(* Logix 5000 project; controller MV vendor 1 type 14 code 217 rev 31.11; software revision 31.00; part 51 of 53 *)
(* tags used below, declared in another part *)
   Alarm_Reset : BOOL;
   CWD : CHECKWORD_FLAGS;
   Default_Check_Time : DINT;
   Item_Faults_Are_Latched : BOOL;
   Item_Simulation_Flag : BOOL;
   MV_MV10R : PlantItem;   // MV10R
   MV_MV10R_ALARM : ALARM_DIGITAL;
   MV_MV10R_D : ALIAS FOR Remote_IO:13:O.Data.9;   // Rouser drive MV10
   MV_MV10R_R : ALIAS FOR Remote_IO:15:I.Data.9;   // MV10 Rouser running signal
   MV_MV11R : PlantItem;   // MV11R
   MV_MV11R_ALARM : ALARM_DIGITAL;
   MV_MV11R_D : ALIAS FOR Remote_IO:13:O.Data.10;   // Rouser drive MV11
   MV_MV11R_R : ALIAS FOR Remote_IO:15:I.Data.10;   // MV11 Rouser running signal
   MV_MV12R : PlantItem;   // MV12R
   MV_MV12R_ALARM : ALARM_DIGITAL;
   MV_MV12R_D : ALIAS FOR Remote_IO:13:O.Data.11;   // Rouser drive MV12
   MV_MV12R_R : ALIAS FOR Remote_IO:15:I.Data.11;   // MV12 Rouser running signal
   MV_MV13R : PlantItem;   // MV13R
   MV_MV13R_ALARM : ALARM_DIGITAL;
   MV_MV13R_D : ALIAS FOR Remote_IO:13:O.Data.12;   // Rouser drive MV13
   MV_MV13R_R : ALIAS FOR Remote_IO:15:I.Data.12;   // MV13 Rouser running signal
   MV_MV14R : PlantItem;   // MV14R
   MV_MV14R_ALARM : ALARM_DIGITAL;
   MV_MV14R_D : ALIAS FOR Remote_IO:13:O.Data.13;   // Rouser drive MV14
   MV_MV14R_R : ALIAS FOR Remote_IO:15:I.Data.13;   // MV14 Rouser running signal
   MV_MV15R : PlantItem;   // MV15R
   MV_MV15R_ALARM : ALARM_DIGITAL;
   MV_MV15R_D : ALIAS FOR Remote_IO:13:O.Data.14;   // Rouser drive MV15
   MV_MV15R_R : ALIAS FOR Remote_IO:15:I.Data.14;   // MV15 Rouser running signal
   MV_MV16R : PlantItem;   // MV16R
   MV_MV16R_ALARM : ALARM_DIGITAL;
   MV_MV16R_D : ALIAS FOR Remote_IO:13:O.Data.15;   // Rouser drive MV16
   MV_MV16R_R : ALIAS FOR Remote_IO:15:I.Data.15;   // MV16 Rouser running signal
   MV_MV17R : PlantItem;   // MV17R
   MV_MV17R_ALARM : ALARM_DIGITAL;
   MV_MV17R_D : ALIAS FOR Remote_IO:14:O.Data.0;   // Rouser drive MV17
   MV_MV17R_R : ALIAS FOR Remote_IO:15:I.Data.16;   // MV17 Rouser running signal
   MV_MV18R : PlantItem;   // MV18R
   MV_MV18R_ALARM : ALARM_DIGITAL;
   MV_MV18R_D : ALIAS FOR Remote_IO:14:O.Data.1;
   MV_MV18R_R : ALIAS FOR Remote_IO:15:I.Data.17;   // MV18 Rouser running signal
   MV_MV19R : PlantItem;   // MV19R
   MV_MV19R_ALARM : ALARM_DIGITAL;
   MV_MV19R_D : ALIAS FOR Remote_IO:14:O.Data.2;   // Rouser drive MV19
   MV_MV19R_R : ALIAS FOR Remote_IO:15:I.Data.18;   // MV19 Rouser running signal
   MV_MV1R : PlantItem;   // MV1R
   MV_MV1R_ALARM : ALARM_DIGITAL;
   MV_MV1R_D : ALIAS FOR Remote_IO:13:O.Data.0;   // Rouser drive MV1
   MV_MV1R_R : ALIAS FOR Remote_IO:15:I.Data.0;
   MV_MV2R : PlantItem;   // MV2R
   MV_MV2R_ALARM : ALARM_DIGITAL;
   MV_MV2R_D : ALIAS FOR Remote_IO:13:O.Data.1;
   MV_MV2R_R : ALIAS FOR Remote_IO:15:I.Data.1;   // MV2 Rouser running signal
   MV_MV30R : PlantItem;   // MV30R
   MV_MV30R_ALARM : ALARM_DIGITAL;
   MV_MV30R_D : ALIAS FOR Remote_IO:14:O.Data.3;   // Rouser drive MV30
   MV_MV30R_R : ALIAS FOR Remote_IO:15:I.Data.19;   // MV30 Rouser running signal
   MV_MV31R : PlantItem;   // MV31R
   MV_MV31R_ALARM : ALARM_DIGITAL;
   MV_MV31R_D : ALIAS FOR Remote_IO:14:O.Data.4;   // Rouser drive MV31
   MV_MV31R_R : ALIAS FOR Remote_IO:15:I.Data.20;   // MV31 Rouser running signal
   MV_MV32R : PlantItem;   // MV32R
   MV_MV32R_ALARM : ALARM_DIGITAL;
   MV_MV32R_D : ALIAS FOR Remote_IO:14:O.Data.5;   // Rouser drive MV32
   MV_MV32R_R : ALIAS FOR Remote_IO:15:I.Data.21;   // MV32 Rouser running signal
   MV_MV33R : PlantItem;   // MV33R
   MV_MV33R_ALARM : ALARM_DIGITAL;
   MV_MV33R_D : ALIAS FOR Remote_IO:14:O.Data.6;   // Rouser drive MV33
   MV_MV33R_R : ALIAS FOR Remote_IO:15:I.Data.22;   // MV33 Rouser running signal
   MV_MV34R : PlantItem;   // MV34R
   MV_MV34R_ALARM : ALARM_DIGITAL;
   MV_MV34R_D : ALIAS FOR Remote_IO:14:O.Data.7;   // Rouser drive MV34
   MV_MV34R_R : ALIAS FOR Remote_IO:15:I.Data.23;   // MV34 Rouser running signal
   MV_MV3R : PlantItem;   // MV3R
   MV_MV3R_ALARM : ALARM_DIGITAL;
   MV_MV3R_D : ALIAS FOR Remote_IO:13:O.Data.2;   // Rouser drive MV3
   MV_MV3R_R : ALIAS FOR Remote_IO:15:I.Data.2;   // MV3 Rouser running signal
   MV_MV4R : PlantItem;   // MV4R
   MV_MV4R_ALARM : ALARM_DIGITAL;
   MV_MV4R_D : ALIAS FOR Remote_IO:13:O.Data.3;   // Rouser drive MV4
   MV_MV4R_R : ALIAS FOR Remote_IO:15:I.Data.3;   // MV4 Rouser running signal
   MV_MV5R : PlantItem;   // MV5R
   MV_MV5R_ALARM : ALARM_DIGITAL;
   MV_MV5R_D : ALIAS FOR Remote_IO:13:O.Data.4;   // Rouser drive MV5
   MV_MV5R_R : ALIAS FOR Remote_IO:15:I.Data.4;   // MV5 Rouser running signal
   MV_MV6R : PlantItem;   // MV6R
   MV_MV6R_ALARM : ALARM_DIGITAL;
   MV_MV6R_D : ALIAS FOR Remote_IO:13:O.Data.5;   // Rouser drive MV6
   MV_MV6R_R : ALIAS FOR Remote_IO:15:I.Data.5;   // MV6 Rouser running signal
   MV_MV7R : PlantItem;   // MV7R
   MV_MV7R_ALARM : ALARM_DIGITAL;
   MV_MV7R_D : ALIAS FOR Remote_IO:13:O.Data.6;   // Rouser drive MV7
   MV_MV7R_R : ALIAS FOR Remote_IO:15:I.Data.6;   // MV7 Rouser running signal
   MV_MV8R : PlantItem;   // MV8R
   MV_MV8R_ALARM : ALARM_DIGITAL;
   MV_MV8R_D : ALIAS FOR Remote_IO:13:O.Data.7;   // Rouser drive MV8
   MV_MV8R_R : ALIAS FOR Remote_IO:15:I.Data.7;   // MV8 Rouser running signal
   MV_MV9R : PlantItem;   // MV9R
   MV_MV9R_ALARM : ALARM_DIGITAL;
   MV_MV9R_D : ALIAS FOR Remote_IO:13:O.Data.8;   // Rouser drive MV9
   MV_MV9R_R : ALIAS FOR Remote_IO:15:I.Data.8;   // MV9 Rouser running signal
   One_Second_One_Scan : ALIAS FOR One_Second_1_scan;
   Scada_Pump_Fault_No : DINT;
   Scada_Pump_H_Fault_No : DINT;
   Scada_Pump_T_Fault_No : DINT;
   Unused_Healthy_Feedback : BOOL;
   Unused_NotTripped_Feedback : BOOL;
(* MV_Common, continued *)

ROUTINE MV_Pumps   (* ladder *)
   0: [NEQ(MV_MV1R.DriveBits,0) OTE(MV_MV1R.CW.[CWD.AUTODRV]) ,[XIC(MV_MV1R.CW.[CWD.AUTODRV]) XIO(MV_MV1R.CW.[CWD.MANUAL]) ,XIC(MV_MV1R.CW.[CWD.MANDRV]) XIC(MV_MV1R.CW.[CWD.MANUAL]) ] OTE(MV_MV1R.CW.[CWD.OUTPUT]) ,XIC(MV_MV1R.CW.[CWD.OUTPUT]) OTE(MV_MV1R_D) ,XIC(S:FS) [OTU(MV_MV1R.CW.[CWD.MANUAL]) ,LEQ(MV_MV1R.CheckTime,0) MOV(Default_Check_Time,MV_MV1R.CheckTime) ] ,[[XIC(MV_MV1R_R) XIO(Item_Simulation_Flag) ,XIC(Item_Simulation_Flag) [XIC(MV_MV1R.CW.[CWD.OUTPUT]) XIO(MV_MV1R.CW.[CWD.SIMFAIL]) ,XIO(MV_MV1R.CW.[CWD.OUTPUT]) XIC(MV_MV1R.CW.[CWD.SIMFAIL]) ] ] OTE(MV_MV1R.CW.[CWD.RUNFB]) ,[XIC(Item_Simulation_Flag) ,XIC(MV_MV1R.CW.[CWD.CHECKOFF]) ,XIC(Unused_Healthy_Feedback) ] OTE(MV_MV1R.CW.[CWD.HEALTHYFB]) ,[XIC(Item_Simulation_Flag) ,XIC(MV_MV1R.CW.[CWD.CHECKOFF]) ,XIC(Unused_NotTripped_Feedback) ] OTE(MV_MV1R.CW.[CWD.NOTTRIPPEDFB]) ] ,[XIC(MV_MV1R.CW.[CWD.AUTODRV]) XIO(MV_MV1R.CW.[CWD.PREVSCAN]) ,XIO(MV_MV1R.CW.[CWD.AUTODRV]) XIC(MV_MV1R.CW.[CWD.PREVSCAN]) ] CLR(MV_MV1R.CheckTimer) ,XIC(One_Second_One_Scan) LES(MV_MV1R.CheckTimer,MV_MV1R.CheckTime) ADD(MV_MV1R.CheckTimer,1,MV_MV1R.CheckTimer) ,XIO(MV_MV1R.CW.[CWD.FAULT]) OTU(MV_MV1R.CW.[CWD.FAULTLOGGED]) ,[GEQ(MV_MV1R.CheckTimer,MV_MV1R.CheckTime) [XIC(MV_MV1R.CW.[CWD.OUTPUT]) XIO(MV_MV1R.CW.[CWD.RUNFB]) ,XIO(MV_MV1R.CW.[CWD.OUTPUT]) XIC(MV_MV1R.CW.[CWD.RUNFB]) ] ,XIO(MV_MV1R.CW.[CWD.HEALTHYFB]) ,XIO(MV_MV1R.CW.[CWD.NOTTRIPPEDFB]) ,XIC(MV_MV1R.CW.[CWD.FAULT]) XIC(Item_Faults_Are_Latched) ,XIC(MV_MV1R.CW.[CWD.HIGHLIGHT]) ] XIO(MV_MV1R.CW.[CWD.CHECKOFF]) XIO(Alarm_Reset) [OTE(MV_MV1R.CW.[CWD.FAULT]) ,ALMD(MV_MV1R_ALARM,0,0,0,0) ] ,XIC(MV_MV1R.CW.[CWD.OUTPUT]) OTE(MV_MV1R.CW.[CWD.PREVSCAN]) ,XIC(MV_MV1R.CW.[CWD.FAULT]) EQU(Scada_Pump_Fault_No,0) XIO(MV_MV1R.CW.[CWD.FAULTLOGGED]) [MOV(20001,Scada_Pump_Fault_No) ,OTL(MV_MV1R.CW.[CWD.FAULTLOGGED]) ] ,XIO(MV_MV1R.CW.[CWD.HEALTHYFB]) EQU(Scada_Pump_H_Fault_No,0) XIO(MV_MV1R.CW.[CWD.HEALTHYFAULTLOGGED]) [MOV(20001,Scada_Pump_H_Fault_No) ,OTL(MV_MV1R.CW.[CWD.HEALTHYFAULTLOGGED]) ] ,XIO(MV_MV1R.CW.[CWD.NOTTRIPPEDFB]) EQU(Scada_Pump_H_Fault_No,0) XIO(MV_MV1R.CW.[CWD.TRIPPEDFAULTLOGGED]) [MOV(20001,Scada_Pump_T_Fault_No) ,OTL(MV_MV1R.CW.[CWD.TRIPPEDFAULTLOGGED]) ] ];
   1: [NEQ(MV_MV2R.DriveBits,0) OTE(MV_MV2R.CW.[CWD.AUTODRV]) ,[XIC(MV_MV2R.CW.[CWD.AUTODRV]) XIO(MV_MV2R.CW.[CWD.MANUAL]) ,XIC(MV_MV2R.CW.[CWD.MANDRV]) XIC(MV_MV2R.CW.[CWD.MANUAL]) ] OTE(MV_MV2R.CW.[CWD.OUTPUT]) ,XIC(MV_MV2R.CW.[CWD.OUTPUT]) OTE(MV_MV2R_D) ,XIC(S:FS) [OTU(MV_MV2R.CW.[CWD.MANUAL]) ,LEQ(MV_MV2R.CheckTime,0) MOV(Default_Check_Time,MV_MV2R.CheckTime) ] ,[[XIC(MV_MV2R_R) XIO(Item_Simulation_Flag) ,XIC(Item_Simulation_Flag) [XIC(MV_MV2R.CW.[CWD.OUTPUT]) XIO(MV_MV2R.CW.[CWD.SIMFAIL]) ,XIO(MV_MV2R.CW.[CWD.OUTPUT]) XIC(MV_MV2R.CW.[CWD.SIMFAIL]) ] ] OTE(MV_MV2R.CW.[CWD.RUNFB]) ,[XIC(Item_Simulation_Flag) ,XIC(MV_MV2R.CW.[CWD.CHECKOFF]) ,XIC(Unused_Healthy_Feedback) ] OTE(MV_MV2R.CW.[CWD.HEALTHYFB]) ,[XIC(Item_Simulation_Flag) ,XIC(MV_MV2R.CW.[CWD.CHECKOFF]) ,XIC(Unused_NotTripped_Feedback) ] OTE(MV_MV2R.CW.[CWD.NOTTRIPPEDFB]) ] ,[XIC(MV_MV2R.CW.[CWD.AUTODRV]) XIO(MV_MV2R.CW.[CWD.PREVSCAN]) ,XIO(MV_MV2R.CW.[CWD.AUTODRV]) XIC(MV_MV2R.CW.[CWD.PREVSCAN]) ] CLR(MV_MV2R.CheckTimer) ,XIC(One_Second_One_Scan) LES(MV_MV2R.CheckTimer,MV_MV2R.CheckTime) ADD(MV_MV2R.CheckTimer,1,MV_MV2R.CheckTimer) ,XIO(MV_MV2R.CW.[CWD.FAULT]) OTU(MV_MV2R.CW.[CWD.FAULTLOGGED]) ,[GEQ(MV_MV2R.CheckTimer,MV_MV2R.CheckTime) [XIC(MV_MV2R.CW.[CWD.OUTPUT]) XIO(MV_MV2R.CW.[CWD.RUNFB]) ,XIO(MV_MV2R.CW.[CWD.OUTPUT]) XIC(MV_MV2R.CW.[CWD.RUNFB]) ] ,XIO(MV_MV2R.CW.[CWD.HEALTHYFB]) ,XIO(MV_MV2R.CW.[CWD.NOTTRIPPEDFB]) ,XIC(MV_MV2R.CW.[CWD.FAULT]) XIC(Item_Faults_Are_Latched) ,XIC(MV_MV2R.CW.[CWD.HIGHLIGHT]) ] XIO(MV_MV2R.CW.[CWD.CHECKOFF]) XIO(Alarm_Reset) [OTE(MV_MV2R.CW.[CWD.FAULT]) ,ALMD(MV_MV2R_ALARM,0,0,0,0) ] ,XIC(MV_MV2R.CW.[CWD.OUTPUT]) OTE(MV_MV2R.CW.[CWD.PREVSCAN]) ,XIC(MV_MV2R.CW.[CWD.FAULT]) EQU(Scada_Pump_Fault_No,0) XIO(MV_MV2R.CW.[CWD.FAULTLOGGED]) [MOV(20001,Scada_Pump_Fault_No) ,OTL(MV_MV2R.CW.[CWD.FAULTLOGGED]) ] ,XIO(MV_MV2R.CW.[CWD.HEALTHYFB]) EQU(Scada_Pump_H_Fault_No,0) XIO(MV_MV2R.CW.[CWD.HEALTHYFAULTLOGGED]) [MOV(20001,Scada_Pump_H_Fault_No) ,OTL(MV_MV2R.CW.[CWD.HEALTHYFAULTLOGGED]) ] ,XIO(MV_MV2R.CW.[CWD.NOTTRIPPEDFB]) EQU(Scada_Pump_H_Fault_No,0) XIO(MV_MV2R.CW.[CWD.TRIPPEDFAULTLOGGED]) [MOV(20001,Scada_Pump_T_Fault_No) ,OTL(MV_MV2R.CW.[CWD.TRIPPEDFAULTLOGGED]) ] ];
   2: [NEQ(MV_MV3R.DriveBits,0) OTE(MV_MV3R.CW.[CWD.AUTODRV]) ,[XIC(MV_MV3R.CW.[CWD.AUTODRV]) XIO(MV_MV3R.CW.[CWD.MANUAL]) ,XIC(MV_MV3R.CW.[CWD.MANDRV]) XIC(MV_MV3R.CW.[CWD.MANUAL]) ] OTE(MV_MV3R.CW.[CWD.OUTPUT]) ,XIC(MV_MV3R.CW.[CWD.OUTPUT]) OTE(MV_MV3R_D) ,XIC(S:FS) [OTU(MV_MV3R.CW.[CWD.MANUAL]) ,LEQ(MV_MV3R.CheckTime,0) MOV(Default_Check_Time,MV_MV3R.CheckTime) ] ,[[XIC(MV_MV3R_R) XIO(Item_Simulation_Flag) ,XIC(Item_Simulation_Flag) [XIC(MV_MV3R.CW.[CWD.OUTPUT]) XIO(MV_MV3R.CW.[CWD.SIMFAIL]) ,XIO(MV_MV3R.CW.[CWD.OUTPUT]) XIC(MV_MV3R.CW.[CWD.SIMFAIL]) ] ] OTE(MV_MV3R.CW.[CWD.RUNFB]) ,[XIC(Item_Simulation_Flag) ,XIC(MV_MV3R.CW.[CWD.CHECKOFF]) ,XIC(Unused_Healthy_Feedback) ] OTE(MV_MV3R.CW.[CWD.HEALTHYFB]) ,[XIC(Item_Simulation_Flag) ,XIC(MV_MV3R.CW.[CWD.CHECKOFF]) ,XIC(Unused_NotTripped_Feedback) ] OTE(MV_MV3R.CW.[CWD.NOTTRIPPEDFB]) ] ,[XIC(MV_MV3R.CW.[CWD.AUTODRV]) XIO(MV_MV3R.CW.[CWD.PREVSCAN]) ,XIO(MV_MV3R.CW.[CWD.AUTODRV]) XIC(MV_MV3R.CW.[CWD.PREVSCAN]) ] CLR(MV_MV3R.CheckTimer) ,XIC(One_Second_One_Scan) LES(MV_MV3R.CheckTimer,MV_MV3R.CheckTime) ADD(MV_MV3R.CheckTimer,1,MV_MV3R.CheckTimer) ,XIO(MV_MV3R.CW.[CWD.FAULT]) OTU(MV_MV3R.CW.[CWD.FAULTLOGGED]) ,[GEQ(MV_MV3R.CheckTimer,MV_MV3R.CheckTime) [XIC(MV_MV3R.CW.[CWD.OUTPUT]) XIO(MV_MV3R.CW.[CWD.RUNFB]) ,XIO(MV_MV3R.CW.[CWD.OUTPUT]) XIC(MV_MV3R.CW.[CWD.RUNFB]) ] ,XIO(MV_MV3R.CW.[CWD.HEALTHYFB]) ,XIO(MV_MV3R.CW.[CWD.NOTTRIPPEDFB]) ,XIC(MV_MV3R.CW.[CWD.FAULT]) XIC(Item_Faults_Are_Latched) ,XIC(MV_MV3R.CW.[CWD.HIGHLIGHT]) ] XIO(MV_MV3R.CW.[CWD.CHECKOFF]) XIO(Alarm_Reset) [OTE(MV_MV3R.CW.[CWD.FAULT]) ,ALMD(MV_MV3R_ALARM,0,0,0,0) ] ,XIC(MV_MV3R.CW.[CWD.OUTPUT]) OTE(MV_MV3R.CW.[CWD.PREVSCAN]) ,XIC(MV_MV3R.CW.[CWD.FAULT]) EQU(Scada_Pump_Fault_No,0) XIO(MV_MV3R.CW.[CWD.FAULTLOGGED]) [MOV(20001,Scada_Pump_Fault_No) ,OTL(MV_MV3R.CW.[CWD.FAULTLOGGED]) ] ,XIO(MV_MV3R.CW.[CWD.HEALTHYFB]) EQU(Scada_Pump_H_Fault_No,0) XIO(MV_MV3R.CW.[CWD.HEALTHYFAULTLOGGED]) [MOV(20001,Scada_Pump_H_Fault_No) ,OTL(MV_MV3R.CW.[CWD.HEALTHYFAULTLOGGED]) ] ,XIO(MV_MV3R.CW.[CWD.NOTTRIPPEDFB]) EQU(Scada_Pump_H_Fault_No,0) XIO(MV_MV3R.CW.[CWD.TRIPPEDFAULTLOGGED]) [MOV(20001,Scada_Pump_T_Fault_No) ,OTL(MV_MV3R.CW.[CWD.TRIPPEDFAULTLOGGED]) ] ];
   3: [NEQ(MV_MV4R.DriveBits,0) OTE(MV_MV4R.CW.[CWD.AUTODRV]) ,[XIC(MV_MV4R.CW.[CWD.AUTODRV]) XIO(MV_MV4R.CW.[CWD.MANUAL]) ,XIC(MV_MV4R.CW.[CWD.MANDRV]) XIC(MV_MV4R.CW.[CWD.MANUAL]) ] OTE(MV_MV4R.CW.[CWD.OUTPUT]) ,XIC(MV_MV4R.CW.[CWD.OUTPUT]) OTE(MV_MV4R_D) ,XIC(S:FS) [OTU(MV_MV4R.CW.[CWD.MANUAL]) ,LEQ(MV_MV4R.CheckTime,0) MOV(Default_Check_Time,MV_MV4R.CheckTime) ] ,[[XIC(MV_MV4R_R) XIO(Item_Simulation_Flag) ,XIC(Item_Simulation_Flag) [XIC(MV_MV4R.CW.[CWD.OUTPUT]) XIO(MV_MV4R.CW.[CWD.SIMFAIL]) ,XIO(MV_MV4R.CW.[CWD.OUTPUT]) XIC(MV_MV4R.CW.[CWD.SIMFAIL]) ] ] OTE(MV_MV4R.CW.[CWD.RUNFB]) ,[XIC(Item_Simulation_Flag) ,XIC(MV_MV4R.CW.[CWD.CHECKOFF]) ,XIC(Unused_Healthy_Feedback) ] OTE(MV_MV4R.CW.[CWD.HEALTHYFB]) ,[XIC(Item_Simulation_Flag) ,XIC(MV_MV4R.CW.[CWD.CHECKOFF]) ,XIC(Unused_NotTripped_Feedback) ] OTE(MV_MV4R.CW.[CWD.NOTTRIPPEDFB]) ] ,[XIC(MV_MV4R.CW.[CWD.AUTODRV]) XIO(MV_MV4R.CW.[CWD.PREVSCAN]) ,XIO(MV_MV4R.CW.[CWD.AUTODRV]) XIC(MV_MV4R.CW.[CWD.PREVSCAN]) ] CLR(MV_MV4R.CheckTimer) ,XIC(One_Second_One_Scan) LES(MV_MV4R.CheckTimer,MV_MV4R.CheckTime) ADD(MV_MV4R.CheckTimer,1,MV_MV4R.CheckTimer) ,XIO(MV_MV4R.CW.[CWD.FAULT]) OTU(MV_MV4R.CW.[CWD.FAULTLOGGED]) ,[GEQ(MV_MV4R.CheckTimer,MV_MV4R.CheckTime) [XIC(MV_MV4R.CW.[CWD.OUTPUT]) XIO(MV_MV4R.CW.[CWD.RUNFB]) ,XIO(MV_MV4R.CW.[CWD.OUTPUT]) XIC(MV_MV4R.CW.[CWD.RUNFB]) ] ,XIO(MV_MV4R.CW.[CWD.HEALTHYFB]) ,XIO(MV_MV4R.CW.[CWD.NOTTRIPPEDFB]) ,XIC(MV_MV4R.CW.[CWD.FAULT]) XIC(Item_Faults_Are_Latched) ,XIC(MV_MV4R.CW.[CWD.HIGHLIGHT]) ] XIO(MV_MV4R.CW.[CWD.CHECKOFF]) XIO(Alarm_Reset) [OTE(MV_MV4R.CW.[CWD.FAULT]) ,ALMD(MV_MV4R_ALARM,0,0,0,0) ] ,XIC(MV_MV4R.CW.[CWD.OUTPUT]) OTE(MV_MV4R.CW.[CWD.PREVSCAN]) ,XIC(MV_MV4R.CW.[CWD.FAULT]) EQU(Scada_Pump_Fault_No,0) XIO(MV_MV4R.CW.[CWD.FAULTLOGGED]) [MOV(20001,Scada_Pump_Fault_No) ,OTL(MV_MV4R.CW.[CWD.FAULTLOGGED]) ] ,XIO(MV_MV4R.CW.[CWD.HEALTHYFB]) EQU(Scada_Pump_H_Fault_No,0) XIO(MV_MV4R.CW.[CWD.HEALTHYFAULTLOGGED]) [MOV(20001,Scada_Pump_H_Fault_No) ,OTL(MV_MV4R.CW.[CWD.HEALTHYFAULTLOGGED]) ] ,XIO(MV_MV4R.CW.[CWD.NOTTRIPPEDFB]) EQU(Scada_Pump_H_Fault_No,0) XIO(MV_MV4R.CW.[CWD.TRIPPEDFAULTLOGGED]) [MOV(20001,Scada_Pump_T_Fault_No) ,OTL(MV_MV4R.CW.[CWD.TRIPPEDFAULTLOGGED]) ] ];
   4: [NEQ(MV_MV5R.DriveBits,0) OTE(MV_MV5R.CW.[CWD.AUTODRV]) ,[XIC(MV_MV5R.CW.[CWD.AUTODRV]) XIO(MV_MV5R.CW.[CWD.MANUAL]) ,XIC(MV_MV5R.CW.[CWD.MANDRV]) XIC(MV_MV5R.CW.[CWD.MANUAL]) ] OTE(MV_MV5R.CW.[CWD.OUTPUT]) ,XIC(MV_MV5R.CW.[CWD.OUTPUT]) OTE(MV_MV5R_D) ,XIC(S:FS) [OTU(MV_MV5R.CW.[CWD.MANUAL]) ,LEQ(MV_MV5R.CheckTime,0) MOV(Default_Check_Time,MV_MV5R.CheckTime) ] ,[[XIC(MV_MV5R_R) XIO(Item_Simulation_Flag) ,XIC(Item_Simulation_Flag) [XIC(MV_MV5R.CW.[CWD.OUTPUT]) XIO(MV_MV5R.CW.[CWD.SIMFAIL]) ,XIO(MV_MV5R.CW.[CWD.OUTPUT]) XIC(MV_MV5R.CW.[CWD.SIMFAIL]) ] ] OTE(MV_MV5R.CW.[CWD.RUNFB]) ,[XIC(Item_Simulation_Flag) ,XIC(MV_MV5R.CW.[CWD.CHECKOFF]) ,XIC(Unused_Healthy_Feedback) ] OTE(MV_MV5R.CW.[CWD.HEALTHYFB]) ,[XIC(Item_Simulation_Flag) ,XIC(MV_MV5R.CW.[CWD.CHECKOFF]) ,XIC(Unused_NotTripped_Feedback) ] OTE(MV_MV5R.CW.[CWD.NOTTRIPPEDFB]) ] ,[XIC(MV_MV5R.CW.[CWD.AUTODRV]) XIO(MV_MV5R.CW.[CWD.PREVSCAN]) ,XIO(MV_MV5R.CW.[CWD.AUTODRV]) XIC(MV_MV5R.CW.[CWD.PREVSCAN]) ] CLR(MV_MV5R.CheckTimer) ,XIC(One_Second_One_Scan) LES(MV_MV5R.CheckTimer,MV_MV5R.CheckTime) ADD(MV_MV5R.CheckTimer,1,MV_MV5R.CheckTimer) ,XIO(MV_MV5R.CW.[CWD.FAULT]) OTU(MV_MV5R.CW.[CWD.FAULTLOGGED]) ,[GEQ(MV_MV5R.CheckTimer,MV_MV5R.CheckTime) [XIC(MV_MV5R.CW.[CWD.OUTPUT]) XIO(MV_MV5R.CW.[CWD.RUNFB]) ,XIO(MV_MV5R.CW.[CWD.OUTPUT]) XIC(MV_MV5R.CW.[CWD.RUNFB]) ] ,XIO(MV_MV5R.CW.[CWD.HEALTHYFB]) ,XIO(MV_MV5R.CW.[CWD.NOTTRIPPEDFB]) ,XIC(MV_MV5R.CW.[CWD.FAULT]) XIC(Item_Faults_Are_Latched) ,XIC(MV_MV5R.CW.[CWD.HIGHLIGHT]) ] XIO(MV_MV5R.CW.[CWD.CHECKOFF]) XIO(Alarm_Reset) [OTE(MV_MV5R.CW.[CWD.FAULT]) ,ALMD(MV_MV5R_ALARM,0,0,0,0) ] ,XIC(MV_MV5R.CW.[CWD.OUTPUT]) OTE(MV_MV5R.CW.[CWD.PREVSCAN]) ,XIC(MV_MV5R.CW.[CWD.FAULT]) EQU(Scada_Pump_Fault_No,0) XIO(MV_MV5R.CW.[CWD.FAULTLOGGED]) [MOV(20001,Scada_Pump_Fault_No) ,OTL(MV_MV5R.CW.[CWD.FAULTLOGGED]) ] ,XIO(MV_MV5R.CW.[CWD.HEALTHYFB]) EQU(Scada_Pump_H_Fault_No,0) XIO(MV_MV5R.CW.[CWD.HEALTHYFAULTLOGGED]) [MOV(20001,Scada_Pump_H_Fault_No) ,OTL(MV_MV5R.CW.[CWD.HEALTHYFAULTLOGGED]) ] ,XIO(MV_MV5R.CW.[CWD.NOTTRIPPEDFB]) EQU(Scada_Pump_H_Fault_No,0) XIO(MV_MV5R.CW.[CWD.TRIPPEDFAULTLOGGED]) [MOV(20001,Scada_Pump_T_Fault_No) ,OTL(MV_MV5R.CW.[CWD.TRIPPEDFAULTLOGGED]) ] ];
   5: [NEQ(MV_MV6R.DriveBits,0) OTE(MV_MV6R.CW.[CWD.AUTODRV]) ,[XIC(MV_MV6R.CW.[CWD.AUTODRV]) XIO(MV_MV6R.CW.[CWD.MANUAL]) ,XIC(MV_MV6R.CW.[CWD.MANDRV]) XIC(MV_MV6R.CW.[CWD.MANUAL]) ] OTE(MV_MV6R.CW.[CWD.OUTPUT]) ,XIC(MV_MV6R.CW.[CWD.OUTPUT]) OTE(MV_MV6R_D) ,XIC(S:FS) [OTU(MV_MV6R.CW.[CWD.MANUAL]) ,LEQ(MV_MV6R.CheckTime,0) MOV(Default_Check_Time,MV_MV6R.CheckTime) ] ,[[XIC(MV_MV6R_R) XIO(Item_Simulation_Flag) ,XIC(Item_Simulation_Flag) [XIC(MV_MV6R.CW.[CWD.OUTPUT]) XIO(MV_MV6R.CW.[CWD.SIMFAIL]) ,XIO(MV_MV6R.CW.[CWD.OUTPUT]) XIC(MV_MV6R.CW.[CWD.SIMFAIL]) ] ] OTE(MV_MV6R.CW.[CWD.RUNFB]) ,[XIC(Item_Simulation_Flag) ,XIC(MV_MV6R.CW.[CWD.CHECKOFF]) ,XIC(Unused_Healthy_Feedback) ] OTE(MV_MV6R.CW.[CWD.HEALTHYFB]) ,[XIC(Item_Simulation_Flag) ,XIC(MV_MV6R.CW.[CWD.CHECKOFF]) ,XIC(Unused_NotTripped_Feedback) ] OTE(MV_MV6R.CW.[CWD.NOTTRIPPEDFB]) ] ,[XIC(MV_MV6R.CW.[CWD.AUTODRV]) XIO(MV_MV6R.CW.[CWD.PREVSCAN]) ,XIO(MV_MV6R.CW.[CWD.AUTODRV]) XIC(MV_MV6R.CW.[CWD.PREVSCAN]) ] CLR(MV_MV6R.CheckTimer) ,XIC(One_Second_One_Scan) LES(MV_MV6R.CheckTimer,MV_MV6R.CheckTime) ADD(MV_MV6R.CheckTimer,1,MV_MV6R.CheckTimer) ,XIO(MV_MV6R.CW.[CWD.FAULT]) OTU(MV_MV6R.CW.[CWD.FAULTLOGGED]) ,[GEQ(MV_MV6R.CheckTimer,MV_MV6R.CheckTime) [XIC(MV_MV6R.CW.[CWD.OUTPUT]) XIO(MV_MV6R.CW.[CWD.RUNFB]) ,XIO(MV_MV6R.CW.[CWD.OUTPUT]) XIC(MV_MV6R.CW.[CWD.RUNFB]) ] ,XIO(MV_MV6R.CW.[CWD.HEALTHYFB]) ,XIO(MV_MV6R.CW.[CWD.NOTTRIPPEDFB]) ,XIC(MV_MV6R.CW.[CWD.FAULT]) XIC(Item_Faults_Are_Latched) ,XIC(MV_MV6R.CW.[CWD.HIGHLIGHT]) ] XIO(MV_MV6R.CW.[CWD.CHECKOFF]) XIO(Alarm_Reset) [OTE(MV_MV6R.CW.[CWD.FAULT]) ,ALMD(MV_MV6R_ALARM,0,0,0,0) ] ,XIC(MV_MV6R.CW.[CWD.OUTPUT]) OTE(MV_MV6R.CW.[CWD.PREVSCAN]) ,XIC(MV_MV6R.CW.[CWD.FAULT]) EQU(Scada_Pump_Fault_No,0) XIO(MV_MV6R.CW.[CWD.FAULTLOGGED]) [MOV(20001,Scada_Pump_Fault_No) ,OTL(MV_MV6R.CW.[CWD.FAULTLOGGED]) ] ,XIO(MV_MV6R.CW.[CWD.HEALTHYFB]) EQU(Scada_Pump_H_Fault_No,0) XIO(MV_MV6R.CW.[CWD.HEALTHYFAULTLOGGED]) [MOV(20001,Scada_Pump_H_Fault_No) ,OTL(MV_MV6R.CW.[CWD.HEALTHYFAULTLOGGED]) ] ,XIO(MV_MV6R.CW.[CWD.NOTTRIPPEDFB]) EQU(Scada_Pump_H_Fault_No,0) XIO(MV_MV6R.CW.[CWD.TRIPPEDFAULTLOGGED]) [MOV(20001,Scada_Pump_T_Fault_No) ,OTL(MV_MV6R.CW.[CWD.TRIPPEDFAULTLOGGED]) ] ];
   6: [NEQ(MV_MV7R.DriveBits,0) OTE(MV_MV7R.CW.[CWD.AUTODRV]) ,[XIC(MV_MV7R.CW.[CWD.AUTODRV]) XIO(MV_MV7R.CW.[CWD.MANUAL]) ,XIC(MV_MV7R.CW.[CWD.MANDRV]) XIC(MV_MV7R.CW.[CWD.MANUAL]) ] OTE(MV_MV7R.CW.[CWD.OUTPUT]) ,XIC(MV_MV7R.CW.[CWD.OUTPUT]) OTE(MV_MV7R_D) ,XIC(S:FS) [OTU(MV_MV7R.CW.[CWD.MANUAL]) ,LEQ(MV_MV7R.CheckTime,0) MOV(Default_Check_Time,MV_MV7R.CheckTime) ] ,[[XIC(MV_MV7R_R) XIO(Item_Simulation_Flag) ,XIC(Item_Simulation_Flag) [XIC(MV_MV7R.CW.[CWD.OUTPUT]) XIO(MV_MV7R.CW.[CWD.SIMFAIL]) ,XIO(MV_MV7R.CW.[CWD.OUTPUT]) XIC(MV_MV7R.CW.[CWD.SIMFAIL]) ] ] OTE(MV_MV7R.CW.[CWD.RUNFB]) ,[XIC(Item_Simulation_Flag) ,XIC(MV_MV7R.CW.[CWD.CHECKOFF]) ,XIC(Unused_Healthy_Feedback) ] OTE(MV_MV7R.CW.[CWD.HEALTHYFB]) ,[XIC(Item_Simulation_Flag) ,XIC(MV_MV7R.CW.[CWD.CHECKOFF]) ,XIC(Unused_NotTripped_Feedback) ] OTE(MV_MV7R.CW.[CWD.NOTTRIPPEDFB]) ] ,[XIC(MV_MV7R.CW.[CWD.AUTODRV]) XIO(MV_MV7R.CW.[CWD.PREVSCAN]) ,XIO(MV_MV7R.CW.[CWD.AUTODRV]) XIC(MV_MV7R.CW.[CWD.PREVSCAN]) ] CLR(MV_MV7R.CheckTimer) ,XIC(One_Second_One_Scan) LES(MV_MV7R.CheckTimer,MV_MV7R.CheckTime) ADD(MV_MV7R.CheckTimer,1,MV_MV7R.CheckTimer) ,XIO(MV_MV7R.CW.[CWD.FAULT]) OTU(MV_MV7R.CW.[CWD.FAULTLOGGED]) ,[GEQ(MV_MV7R.CheckTimer,MV_MV7R.CheckTime) [XIC(MV_MV7R.CW.[CWD.OUTPUT]) XIO(MV_MV7R.CW.[CWD.RUNFB]) ,XIO(MV_MV7R.CW.[CWD.OUTPUT]) XIC(MV_MV7R.CW.[CWD.RUNFB]) ] ,XIO(MV_MV7R.CW.[CWD.HEALTHYFB]) ,XIO(MV_MV7R.CW.[CWD.NOTTRIPPEDFB]) ,XIC(MV_MV7R.CW.[CWD.FAULT]) XIC(Item_Faults_Are_Latched) ,XIC(MV_MV7R.CW.[CWD.HIGHLIGHT]) ] XIO(MV_MV7R.CW.[CWD.CHECKOFF]) XIO(Alarm_Reset) [OTE(MV_MV7R.CW.[CWD.FAULT]) ,ALMD(MV_MV7R_ALARM,0,0,0,0) ] ,XIC(MV_MV7R.CW.[CWD.OUTPUT]) OTE(MV_MV7R.CW.[CWD.PREVSCAN]) ,XIC(MV_MV7R.CW.[CWD.FAULT]) EQU(Scada_Pump_Fault_No,0) XIO(MV_MV7R.CW.[CWD.FAULTLOGGED]) [MOV(20001,Scada_Pump_Fault_No) ,OTL(MV_MV7R.CW.[CWD.FAULTLOGGED]) ] ,XIO(MV_MV7R.CW.[CWD.HEALTHYFB]) EQU(Scada_Pump_H_Fault_No,0) XIO(MV_MV7R.CW.[CWD.HEALTHYFAULTLOGGED]) [MOV(20001,Scada_Pump_H_Fault_No) ,OTL(MV_MV7R.CW.[CWD.HEALTHYFAULTLOGGED]) ] ,XIO(MV_MV7R.CW.[CWD.NOTTRIPPEDFB]) EQU(Scada_Pump_H_Fault_No,0) XIO(MV_MV7R.CW.[CWD.TRIPPEDFAULTLOGGED]) [MOV(20001,Scada_Pump_T_Fault_No) ,OTL(MV_MV7R.CW.[CWD.TRIPPEDFAULTLOGGED]) ] ];
   7: [NEQ(MV_MV8R.DriveBits,0) OTE(MV_MV8R.CW.[CWD.AUTODRV]) ,[XIC(MV_MV8R.CW.[CWD.AUTODRV]) XIO(MV_MV8R.CW.[CWD.MANUAL]) ,XIC(MV_MV8R.CW.[CWD.MANDRV]) XIC(MV_MV8R.CW.[CWD.MANUAL]) ] OTE(MV_MV8R.CW.[CWD.OUTPUT]) ,XIC(MV_MV8R.CW.[CWD.OUTPUT]) OTE(MV_MV8R_D) ,XIC(S:FS) [OTU(MV_MV8R.CW.[CWD.MANUAL]) ,LEQ(MV_MV8R.CheckTime,0) MOV(Default_Check_Time,MV_MV8R.CheckTime) ] ,[[XIC(MV_MV8R_R) XIO(Item_Simulation_Flag) ,XIC(Item_Simulation_Flag) [XIC(MV_MV8R.CW.[CWD.OUTPUT]) XIO(MV_MV8R.CW.[CWD.SIMFAIL]) ,XIO(MV_MV8R.CW.[CWD.OUTPUT]) XIC(MV_MV8R.CW.[CWD.SIMFAIL]) ] ] OTE(MV_MV8R.CW.[CWD.RUNFB]) ,[XIC(Item_Simulation_Flag) ,XIC(MV_MV8R.CW.[CWD.CHECKOFF]) ,XIC(Unused_Healthy_Feedback) ] OTE(MV_MV8R.CW.[CWD.HEALTHYFB]) ,[XIC(Item_Simulation_Flag) ,XIC(MV_MV8R.CW.[CWD.CHECKOFF]) ,XIC(Unused_NotTripped_Feedback) ] OTE(MV_MV8R.CW.[CWD.NOTTRIPPEDFB]) ] ,[XIC(MV_MV8R.CW.[CWD.AUTODRV]) XIO(MV_MV8R.CW.[CWD.PREVSCAN]) ,XIO(MV_MV8R.CW.[CWD.AUTODRV]) XIC(MV_MV8R.CW.[CWD.PREVSCAN]) ] CLR(MV_MV8R.CheckTimer) ,XIC(One_Second_One_Scan) LES(MV_MV8R.CheckTimer,MV_MV8R.CheckTime) ADD(MV_MV8R.CheckTimer,1,MV_MV8R.CheckTimer) ,XIO(MV_MV8R.CW.[CWD.FAULT]) OTU(MV_MV8R.CW.[CWD.FAULTLOGGED]) ,[GEQ(MV_MV8R.CheckTimer,MV_MV8R.CheckTime) [XIC(MV_MV8R.CW.[CWD.OUTPUT]) XIO(MV_MV8R.CW.[CWD.RUNFB]) ,XIO(MV_MV8R.CW.[CWD.OUTPUT]) XIC(MV_MV8R.CW.[CWD.RUNFB]) ] ,XIO(MV_MV8R.CW.[CWD.HEALTHYFB]) ,XIO(MV_MV8R.CW.[CWD.NOTTRIPPEDFB]) ,XIC(MV_MV8R.CW.[CWD.FAULT]) XIC(Item_Faults_Are_Latched) ,XIC(MV_MV8R.CW.[CWD.HIGHLIGHT]) ] XIO(MV_MV8R.CW.[CWD.CHECKOFF]) XIO(Alarm_Reset) [OTE(MV_MV8R.CW.[CWD.FAULT]) ,ALMD(MV_MV8R_ALARM,0,0,0,0) ] ,XIC(MV_MV8R.CW.[CWD.OUTPUT]) OTE(MV_MV8R.CW.[CWD.PREVSCAN]) ,XIC(MV_MV8R.CW.[CWD.FAULT]) EQU(Scada_Pump_Fault_No,0) XIO(MV_MV8R.CW.[CWD.FAULTLOGGED]) [MOV(20001,Scada_Pump_Fault_No) ,OTL(MV_MV8R.CW.[CWD.FAULTLOGGED]) ] ,XIO(MV_MV8R.CW.[CWD.HEALTHYFB]) EQU(Scada_Pump_H_Fault_No,0) XIO(MV_MV8R.CW.[CWD.HEALTHYFAULTLOGGED]) [MOV(20001,Scada_Pump_H_Fault_No) ,OTL(MV_MV8R.CW.[CWD.HEALTHYFAULTLOGGED]) ] ,XIO(MV_MV8R.CW.[CWD.NOTTRIPPEDFB]) EQU(Scada_Pump_H_Fault_No,0) XIO(MV_MV8R.CW.[CWD.TRIPPEDFAULTLOGGED]) [MOV(20001,Scada_Pump_T_Fault_No) ,OTL(MV_MV8R.CW.[CWD.TRIPPEDFAULTLOGGED]) ] ];
   8: [NEQ(MV_MV9R.DriveBits,0) OTE(MV_MV9R.CW.[CWD.AUTODRV]) ,[XIC(MV_MV9R.CW.[CWD.AUTODRV]) XIO(MV_MV9R.CW.[CWD.MANUAL]) ,XIC(MV_MV9R.CW.[CWD.MANDRV]) XIC(MV_MV9R.CW.[CWD.MANUAL]) ] OTE(MV_MV9R.CW.[CWD.OUTPUT]) ,XIC(MV_MV9R.CW.[CWD.OUTPUT]) OTE(MV_MV9R_D) ,XIC(S:FS) [OTU(MV_MV9R.CW.[CWD.MANUAL]) ,LEQ(MV_MV9R.CheckTime,0) MOV(Default_Check_Time,MV_MV9R.CheckTime) ] ,[[XIC(MV_MV9R_R) XIO(Item_Simulation_Flag) ,XIC(Item_Simulation_Flag) [XIC(MV_MV9R.CW.[CWD.OUTPUT]) XIO(MV_MV9R.CW.[CWD.SIMFAIL]) ,XIO(MV_MV9R.CW.[CWD.OUTPUT]) XIC(MV_MV9R.CW.[CWD.SIMFAIL]) ] ] OTE(MV_MV9R.CW.[CWD.RUNFB]) ,[XIC(Item_Simulation_Flag) ,XIC(MV_MV9R.CW.[CWD.CHECKOFF]) ,XIC(Unused_Healthy_Feedback) ] OTE(MV_MV9R.CW.[CWD.HEALTHYFB]) ,[XIC(Item_Simulation_Flag) ,XIC(MV_MV9R.CW.[CWD.CHECKOFF]) ,XIC(Unused_NotTripped_Feedback) ] OTE(MV_MV9R.CW.[CWD.NOTTRIPPEDFB]) ] ,[XIC(MV_MV9R.CW.[CWD.AUTODRV]) XIO(MV_MV9R.CW.[CWD.PREVSCAN]) ,XIO(MV_MV9R.CW.[CWD.AUTODRV]) XIC(MV_MV9R.CW.[CWD.PREVSCAN]) ] CLR(MV_MV9R.CheckTimer) ,XIC(One_Second_One_Scan) LES(MV_MV9R.CheckTimer,MV_MV9R.CheckTime) ADD(MV_MV9R.CheckTimer,1,MV_MV9R.CheckTimer) ,XIO(MV_MV9R.CW.[CWD.FAULT]) OTU(MV_MV9R.CW.[CWD.FAULTLOGGED]) ,[GEQ(MV_MV9R.CheckTimer,MV_MV9R.CheckTime) [XIC(MV_MV9R.CW.[CWD.OUTPUT]) XIO(MV_MV9R.CW.[CWD.RUNFB]) ,XIO(MV_MV9R.CW.[CWD.OUTPUT]) XIC(MV_MV9R.CW.[CWD.RUNFB]) ] ,XIO(MV_MV9R.CW.[CWD.HEALTHYFB]) ,XIO(MV_MV9R.CW.[CWD.NOTTRIPPEDFB]) ,XIC(MV_MV9R.CW.[CWD.FAULT]) XIC(Item_Faults_Are_Latched) ,XIC(MV_MV9R.CW.[CWD.HIGHLIGHT]) ] XIO(MV_MV9R.CW.[CWD.CHECKOFF]) XIO(Alarm_Reset) [OTE(MV_MV9R.CW.[CWD.FAULT]) ,ALMD(MV_MV9R_ALARM,0,0,0,0) ] ,XIC(MV_MV9R.CW.[CWD.OUTPUT]) OTE(MV_MV9R.CW.[CWD.PREVSCAN]) ,XIC(MV_MV9R.CW.[CWD.FAULT]) EQU(Scada_Pump_Fault_No,0) XIO(MV_MV9R.CW.[CWD.FAULTLOGGED]) [MOV(20001,Scada_Pump_Fault_No) ,OTL(MV_MV9R.CW.[CWD.FAULTLOGGED]) ] ,XIO(MV_MV9R.CW.[CWD.HEALTHYFB]) EQU(Scada_Pump_H_Fault_No,0) XIO(MV_MV9R.CW.[CWD.HEALTHYFAULTLOGGED]) [MOV(20001,Scada_Pump_H_Fault_No) ,OTL(MV_MV9R.CW.[CWD.HEALTHYFAULTLOGGED]) ] ,XIO(MV_MV9R.CW.[CWD.NOTTRIPPEDFB]) EQU(Scada_Pump_H_Fault_No,0) XIO(MV_MV9R.CW.[CWD.TRIPPEDFAULTLOGGED]) [MOV(20001,Scada_Pump_T_Fault_No) ,OTL(MV_MV9R.CW.[CWD.TRIPPEDFAULTLOGGED]) ] ];
   9: [NEQ(MV_MV10R.DriveBits,0) OTE(MV_MV10R.CW.[CWD.AUTODRV]) ,[XIC(MV_MV10R.CW.[CWD.AUTODRV]) XIO(MV_MV10R.CW.[CWD.MANUAL]) ,XIC(MV_MV10R.CW.[CWD.MANDRV]) XIC(MV_MV10R.CW.[CWD.MANUAL]) ] OTE(MV_MV10R.CW.[CWD.OUTPUT]) ,XIC(MV_MV10R.CW.[CWD.OUTPUT]) OTE(MV_MV10R_D) ,XIC(S:FS) [OTU(MV_MV10R.CW.[CWD.MANUAL]) ,LEQ(MV_MV10R.CheckTime,0) MOV(Default_Check_Time,MV_MV10R.CheckTime) ] ,[[XIC(MV_MV10R_R) XIO(Item_Simulation_Flag) ,XIC(Item_Simulation_Flag) [XIC(MV_MV10R.CW.[CWD.OUTPUT]) XIO(MV_MV10R.CW.[CWD.SIMFAIL]) ,XIO(MV_MV10R.CW.[CWD.OUTPUT]) XIC(MV_MV10R.CW.[CWD.SIMFAIL]) ] ] OTE(MV_MV10R.CW.[CWD.RUNFB]) ,[XIC(Item_Simulation_Flag) ,XIC(MV_MV10R.CW.[CWD.CHECKOFF]) ,XIC(Unused_Healthy_Feedback) ] OTE(MV_MV10R.CW.[CWD.HEALTHYFB]) ,[XIC(Item_Simulation_Flag) ,XIC(MV_MV10R.CW.[CWD.CHECKOFF]) ,XIC(Unused_NotTripped_Feedback) ] OTE(MV_MV10R.CW.[CWD.NOTTRIPPEDFB]) ] ,[XIC(MV_MV10R.CW.[CWD.AUTODRV]) XIO(MV_MV10R.CW.[CWD.PREVSCAN]) ,XIO(MV_MV10R.CW.[CWD.AUTODRV]) XIC(MV_MV10R.CW.[CWD.PREVSCAN]) ] CLR(MV_MV10R.CheckTimer) ,XIC(One_Second_One_Scan) LES(MV_MV10R.CheckTimer,MV_MV10R.CheckTime) ADD(MV_MV10R.CheckTimer,1,MV_MV10R.CheckTimer) ,XIO(MV_MV10R.CW.[CWD.FAULT]) OTU(MV_MV10R.CW.[CWD.FAULTLOGGED]) ,[GEQ(MV_MV10R.CheckTimer,MV_MV10R.CheckTime) [XIC(MV_MV10R.CW.[CWD.OUTPUT]) XIO(MV_MV10R.CW.[CWD.RUNFB]) ,XIO(MV_MV10R.CW.[CWD.OUTPUT]) XIC(MV_MV10R.CW.[CWD.RUNFB]) ] ,XIO(MV_MV10R.CW.[CWD.HEALTHYFB]) ,XIO(MV_MV10R.CW.[CWD.NOTTRIPPEDFB]) ,XIC(MV_MV10R.CW.[CWD.FAULT]) XIC(Item_Faults_Are_Latched) ,XIC(MV_MV10R.CW.[CWD.HIGHLIGHT]) ] XIO(MV_MV10R.CW.[CWD.CHECKOFF]) XIO(Alarm_Reset) [OTE(MV_MV10R.CW.[CWD.FAULT]) ,ALMD(MV_MV10R_ALARM,0,0,0,0) ] ,XIC(MV_MV10R.CW.[CWD.OUTPUT]) OTE(MV_MV10R.CW.[CWD.PREVSCAN]) ,XIC(MV_MV10R.CW.[CWD.FAULT]) EQU(Scada_Pump_Fault_No,0) XIO(MV_MV10R.CW.[CWD.FAULTLOGGED]) [MOV(20001,Scada_Pump_Fault_No) ,OTL(MV_MV10R.CW.[CWD.FAULTLOGGED]) ] ,XIO(MV_MV10R.CW.[CWD.HEALTHYFB]) EQU(Scada_Pump_H_Fault_No,0) XIO(MV_MV10R.CW.[CWD.HEALTHYFAULTLOGGED]) [MOV(20001,Scada_Pump_H_Fault_No) ,OTL(MV_MV10R.CW.[CWD.HEALTHYFAULTLOGGED]) ] ,XIO(MV_MV10R.CW.[CWD.NOTTRIPPEDFB]) EQU(Scada_Pump_H_Fault_No,0) XIO(MV_MV10R.CW.[CWD.TRIPPEDFAULTLOGGED]) [MOV(20001,Scada_Pump_T_Fault_No) ,OTL(MV_MV10R.CW.[CWD.TRIPPEDFAULTLOGGED]) ] ];
   10: [NEQ(MV_MV11R.DriveBits,0) OTE(MV_MV11R.CW.[CWD.AUTODRV]) ,[XIC(MV_MV11R.CW.[CWD.AUTODRV]) XIO(MV_MV11R.CW.[CWD.MANUAL]) ,XIC(MV_MV11R.CW.[CWD.MANDRV]) XIC(MV_MV11R.CW.[CWD.MANUAL]) ] OTE(MV_MV11R.CW.[CWD.OUTPUT]) ,XIC(MV_MV11R.CW.[CWD.OUTPUT]) OTE(MV_MV11R_D) ,XIC(S:FS) [OTU(MV_MV11R.CW.[CWD.MANUAL]) ,LEQ(MV_MV11R.CheckTime,0) MOV(Default_Check_Time,MV_MV11R.CheckTime) ] ,[[XIC(MV_MV11R_R) XIO(Item_Simulation_Flag) ,XIC(Item_Simulation_Flag) [XIC(MV_MV11R.CW.[CWD.OUTPUT]) XIO(MV_MV11R.CW.[CWD.SIMFAIL]) ,XIO(MV_MV11R.CW.[CWD.OUTPUT]) XIC(MV_MV11R.CW.[CWD.SIMFAIL]) ] ] OTE(MV_MV11R.CW.[CWD.RUNFB]) ,[XIC(Item_Simulation_Flag) ,XIC(MV_MV11R.CW.[CWD.CHECKOFF]) ,XIC(Unused_Healthy_Feedback) ] OTE(MV_MV11R.CW.[CWD.HEALTHYFB]) ,[XIC(Item_Simulation_Flag) ,XIC(MV_MV11R.CW.[CWD.CHECKOFF]) ,XIC(Unused_NotTripped_Feedback) ] OTE(MV_MV11R.CW.[CWD.NOTTRIPPEDFB]) ] ,[XIC(MV_MV11R.CW.[CWD.AUTODRV]) XIO(MV_MV11R.CW.[CWD.PREVSCAN]) ,XIO(MV_MV11R.CW.[CWD.AUTODRV]) XIC(MV_MV11R.CW.[CWD.PREVSCAN]) ] CLR(MV_MV11R.CheckTimer) ,XIC(One_Second_One_Scan) LES(MV_MV11R.CheckTimer,MV_MV11R.CheckTime) ADD(MV_MV11R.CheckTimer,1,MV_MV11R.CheckTimer) ,XIO(MV_MV11R.CW.[CWD.FAULT]) OTU(MV_MV11R.CW.[CWD.FAULTLOGGED]) ,[GEQ(MV_MV11R.CheckTimer,MV_MV11R.CheckTime) [XIC(MV_MV11R.CW.[CWD.OUTPUT]) XIO(MV_MV11R.CW.[CWD.RUNFB]) ,XIO(MV_MV11R.CW.[CWD.OUTPUT]) XIC(MV_MV11R.CW.[CWD.RUNFB]) ] ,XIO(MV_MV11R.CW.[CWD.HEALTHYFB]) ,XIO(MV_MV11R.CW.[CWD.NOTTRIPPEDFB]) ,XIC(MV_MV11R.CW.[CWD.FAULT]) XIC(Item_Faults_Are_Latched) ,XIC(MV_MV11R.CW.[CWD.HIGHLIGHT]) ] XIO(MV_MV11R.CW.[CWD.CHECKOFF]) XIO(Alarm_Reset) [OTE(MV_MV11R.CW.[CWD.FAULT]) ,ALMD(MV_MV11R_ALARM,0,0,0,0) ] ,XIC(MV_MV11R.CW.[CWD.OUTPUT]) OTE(MV_MV11R.CW.[CWD.PREVSCAN]) ,XIC(MV_MV11R.CW.[CWD.FAULT]) EQU(Scada_Pump_Fault_No,0) XIO(MV_MV11R.CW.[CWD.FAULTLOGGED]) [MOV(20001,Scada_Pump_Fault_No) ,OTL(MV_MV11R.CW.[CWD.FAULTLOGGED]) ] ,XIO(MV_MV11R.CW.[CWD.HEALTHYFB]) EQU(Scada_Pump_H_Fault_No,0) XIO(MV_MV11R.CW.[CWD.HEALTHYFAULTLOGGED]) [MOV(20001,Scada_Pump_H_Fault_No) ,OTL(MV_MV11R.CW.[CWD.HEALTHYFAULTLOGGED]) ] ,XIO(MV_MV11R.CW.[CWD.NOTTRIPPEDFB]) EQU(Scada_Pump_H_Fault_No,0) XIO(MV_MV11R.CW.[CWD.TRIPPEDFAULTLOGGED]) [MOV(20001,Scada_Pump_T_Fault_No) ,OTL(MV_MV11R.CW.[CWD.TRIPPEDFAULTLOGGED]) ] ];